ScreenModuleEditorView "PB: KP8 Stop Runtime (Text Label)" 68x66
   Button "Station Select" at 0,0 size 68x66; TextOff 'STOP RUNTIME'
      Appearance <- "Interface.animate"
*)

(* ===== HMI "HMI_RT_1" =====
system functions are stored by id; their names below are inferred from use

ScreenModuleEditorView "PB: Graphic/Text List" 65x45
   Button "Previous Station Group" at 0,0 size 65x45; TextOff 'Text'
      on Press: SetBit("Interface.actuate")
      Visibility <- "Interface.animate"
      ObjectEnable <- "Interface.animate"
      Appearance <- "Interface.animate"
*)

(* ===== HMI "HMI_RT_1" =====
system functions are stored by id; their names below are inferred from use

ScreenModuleEditorView "PB: Static Text Label" 274x45
   Button "Select All Stations" at 0,0 size 274x45; TextOff 'Text'
      on Press: function_b14e0dd5("Interface.actuate", 0)
      Appearance <- "Interface.animate"
*)

(* ===== HMI "HMI_RT_1" =====
system functions are stored by id; their names below are inferred from use

ScreenModuleEditorView "PB: Static Text Label" 274x45
   Button "Select All Stations" at 0,0 size 274x45; TextOff 'Text'
      on Press: function_b14e0dd5("Interface.actuate", 0)
      Appearance <- "Interface.animate"
*)

(* ===== HMI "HMI_RT_1" =====
system functions are stored by id; their names below are inferred from use

ScreenModuleEditorView "PB: Graphic/Text List" 65x45
   Button "Previous Station Group" at 0,0 size 65x45; TextOff 'Text'
      on Press: SetBit("Interface.actuate")
      Visibility <- "Interface.animate"
      ObjectEnable <- "Interface.animate"
      Appearance <- "Interface.animate"
*)

(* ===== HMI "HMI_RT_1" =====
system functions are stored by id; their names below are inferred from use

ScreenModuleEditorView "PB: Station Select (Text Label)" 205x65
   Button "Station Select" at 0,0 size 205x65; TextOff 'Text'
      on Press: function_b14e0dd5("Interface.actuate", 0)
      Appearance <- "Interface.animate"
*)

(* ===== HMI "HMI_RT_1" =====
system functions are stored by id; their names below are inferred from use

ScreenModuleEditorView "PB: Graphic/Text List" 65x45
   Button "Previous Station Group" at 0,0 size 65x45; TextOff 'Text'
      on Press: function_b14e0dd5("Interface.actuate", 0)
      Visibility <- "Interface.animate"
      ObjectEnable <- "Interface.animate"
      Appearance <- "Interface.animate"
*)

(* ===== HMI "HMI_RT_1" =====
system functions are stored by id; their names below are inferred from use

ScreenModuleEditorView "Drop Zone Label" 240x40
   IOField "Drop Zone Entry" at 171,0 size 69x40; FormatPattern ??
      on OnFinishInput: SetBit("Interface.inputFinished")
      Appearance <- "Interface.animate.ioField"
      ObjectEnable <- "Interface.animate.ioField"
      Visibility <- "Interface.animate.ioField"
      ProcessValue <- "Interface.value"
   TextField "Drop Zone Label" at 0,0 size 240x40; Text 'Drop Zone:'
      Visibility <- "Interface.animate.bg"
      Appearance <- "Interface.animate.bg"
*)

(* ===== HMI "HMI_RT_1" =====
system functions are stored by id; their names below are inferred from use

ScreenModuleEditorView "IO Field: Double Width; Stacked" 414x50
   IOField "PN Entry Field" at 0,0 size 414x50; FormatPattern ????????????????????????????????????????
      on OnFinishInput: SetBit("Interface.inputFinished")
      Appearance <- "Interface.animate"
      ObjectEnable <- "Interface.animate"
      ProcessValue <- "Interface.value"
*)

(* ===== HMI "HMI_RT_1" =====
system functions are stored by id; their names below are inferred from use

ScreenModuleEditorView "IO Field: Timer" 137x50
   IOField "Allotted Time Entry Field" at 0,0 size 137x50; FormatPattern ???????
      on OnFinishInput: SetBit("Interface.inputFinished")
      Appearance <- "Interface.animate"
      ObjectEnable <- "Interface.animate"
      ProcessValue <- "Interface.value"
*)

(* ===== HMI "HMI_RT_1" =====

ScreenModuleEditorView "LED Row" 440x28
   TextField "tfLine" at 0,0 size 110x28; Text 'Text'
      Visibility <- "interface.tfLine.visibility"
      Appearance <- "interface.tfLine.animator"
   TextField "tfTime" at 349,0 size 91x28; Text 'Text'
      Visibility <- "interface.tfTime.visibility"
      Appearance <- "interface.tfTime.animator"
   TextField "tfDropZone" at 105,0 size 42x28; Text 'Text'
      Visibility <- "interface.tfDropZone.visibility"
      Appearance <- "interface.tfDropZone.animator"
   TextField "tfSLPartNumber" at 146,0 size 209x28; Text 'Text'
      Visibility <- "interface.tfPartNumber.count"
      Appearance <- "interface.tfPartNumber.animator"
   TextField "tfDLPartNumber" at 146,0 size 209x28; Text 'Text'
      Visibility <- "interface.tfPartNumber.count"
      Appearance <- "interface.tfPartNumber.animator"
*)

(* ===== HMI "HMI_RT_1" =====
system functions are stored by id; their names below are inferred from use

ScreenModuleEditorView "Line Label" 267x40
   IOField "Line" at 86,0 size 181x40; FormatPattern ?????????
      on OnFinishInput: SetBit("interface.inputFinished")
      Appearance <- "interface.animate.ioField"
      ObjectEnable <- "interface.animate.ioField"
      Visibility <- "interface.animate.ioField"
      ProcessValue <- "interface.value"
   TextField "Line Label" at 0,0 size 267x40; Text 'Line:'
      Visibility <- "interface.animate.bg"
      Appearance <- "interface.animate.bg"
*)

(* ===== HMI "HMI_RT_1" =====
system functions are stored by id; their names below are inferred from use

ScreenModuleEditorView "PB: Graphic/Text List" 65x45
   Button "Previous Station Group" at 0,0 size 65x45; TextOff 'Text'
      on Press: function_b14e0dd5("Interface.actuate", 0)
      Visibility <- "Interface.animate"
      ObjectEnable <- "Interface.animate"
      Appearance <- "Interface.animate"
*)

(* ===== HMI "HMI_RT_1" =====
system functions are stored by id; their names below are inferred from use

ScreenModuleEditorView "PB: KP8 Button Select (Text Label)" 68x66
   Button "Station Select" at 0,0 size 68x66; TextOff 'Text'
      on Press: function_b14e0dd5("Interface.actuate", 0)
      Appearance <- "Interface.animate"
*)

(* ===== HMI "HMI_RT_1" =====

ScreenModuleEditorView "PB: KP8 Reset Button (Text Label" 68x66
   Button "Station Select" at 0,0 size 68x66; TextOff 'RESET SELECTED'
      Appearance <- "Interface.animate"
*)

(* ===== HMI "HMI_RT_1" =====

ScreenModuleEditorView "PB: KP8 Stop Runtime (Text Label)" 68x66
   Button "Station Select" at 0,0 size 68x66; TextOff 'STOP RUNTIME'
      Appearance <- "Interface.animate"
*)

(* ===== HMI "HMI_RT_1" =====
system functions are stored by id; their names below are inferred from use

ScreenModuleEditorView "PB: Station Select (Text Label)" 205x65
   Button "Station Select" at 0,0 size 205x65; TextOff 'Text'
      on Press: function_b14e0dd5("Interface.actuate", 0)
      Appearance <- "Interface.animate"
*)

(* ===== HMI "HMI_RT_1" =====
system functions are stored by id; their names below are inferred from use

ScreenModuleEditorView "PB: Static Text Label" 274x45
   Button "Select All Stations" at 0,0 size 274x45; TextOff 'Text'
      on Press: function_b14e0dd5("Interface.actuate", 0)
      Appearance <- "Interface.animate"
*)

(* ===== HMI "HMI_RT_1" =====
system functions are stored by id; their names below are inferred from use

ScreenModuleEditorView "Station Assignment: Button Details" 513x74
   TextField "Button Label" at 0,0 size 75x74; Text 'Text'
      Visibility <- "Interface.label.animate"
      Appearance <- "Interface.label.animate"
   TextField "Critical Time" at 70,37 size 122x37; Text 'Text'
      Visibility <- "Interface.critical.animate"
      Appearance <- "Interface.critical.animate"
   TextField "Alloted Time" at 70,0 size 122x38; Text 'Text'
      Visibility <- "Interface.alloted.animate"
      Appearance <- "Interface.alloted.animate"
   TextField "Part Number" at 185,0 size 328x74; Text 'Text'
      Visibility <- "Interface.partNumber.animate"
      Appearance <- "Interface.partNumber.animate"
   Button "Select PB" at 0,0 size 513x74; TextOff 'Text'
      on Press: function_b14e0dd5("Interface.select.actuate", 0)
      Visibility <- "Interface.select.animate"
      ObjectEnable <- "Interface.select.animate"
*)

(* ===== HMI "HMI_RT_1" =====
system functions are stored by id; their names below are inferred from use

ScreenModuleEditorView "Table Row" 1312x52
   TextField "tfLine" at 5,1 size 216x48; Text 'Text'
      Visibility <- "interface.tfLine.visibility"
      Appearance <- "interface.tfLine.animator"
   TextField "tfTime" at 1085,1 size 222x48; Text 'Text'
      Visibility <- "interface.tfTime.visibility"
      Appearance <- "interface.tfTime.animator"
   TextField "tfDropZone" at 211,1 size 236x48; Text 'Text'
      Visibility <- "interface.tfDropZone.visibility"
      Appearance <- "interface.tfDropZone.animator"
   TextField "tfSLPartNumber" at 445,1 size 650x48; Text 'Text'
      Visibility <- "interface.tfPartNumber.count"
      Appearance <- "interface.tfPartNumber.animator"
   Button "pbSelect" at 0,0 size 1312x52; TextOff 'Text'
      on Release: ResetBit("interface.pbSelection.request")
      on Press: SetBit("interface.pbSelection.request")
      Visibility <- "interface.pbSelection.visibility"
   Rectangle "rtBackground" at 0,0 size 1312x52
      Visibility <- "interface.rtBackground.visibility"
   TextField "tfDLPartNumber" at 445,1 size 650x48; Text 'Text'
      Visibility <- "interface.tfPartNumber.count"
      Appearance <- "interface.tfPartNumber.animator"
*)

(* ===== HMI "HMI_RT_1" =====
system functions are stored by id; their names below are inferred from use

ScreenModuleEditorView "PB: Static Text Label" 274x45
   Button "Select All Stations" at 0,0 size 274x45; TextOff 'Text'
      on Press: function_b14e0dd5("Interface.actuate", 0)
      Appearance <- "Interface.animate"
      ObjectEnable <- "Interface.animate"
*)

(* ===== HMI "HMI_RT_1" =====
system functions are stored by id; their names below are inferred from use

ScreenModuleEditorView "PB: KP8 Button Select (Text Label)" 68x66
   Button "Station Select" at 0,0 size 68x66; TextOff 'Text'
      on Press: function_b14e0dd5("Interface.actuate", 0)
      Appearance <- "Interface.animate"
      ObjectEnable <- "Interface.animate"
*)

(* ===== HMI "HMI_RT_1" =====
system functions are stored by id; their names below are inferred from use

ScreenModuleEditorView "PB: KP8 Reset Button (Text Label" 68x66
   Button "Station Select" at 0,0 size 68x66; TextOff 'RESET SELECTED'
      Appearance <- "Interface.animate"
      on Press: function_b14e0dd5("Interface.actuate", 0)
*)

(* ===== HMI "HMI_RT_1" =====
system functions are stored by id; their names below are inferred from use

ScreenModuleEditorView "Drop Zone Label" 240x40
   IOField "Drop Zone Entry" at 171,0 size 69x40; FormatPattern ??
      on OnFinishInput: SetBit("Interface.inputFinished")
      Appearance <- "Interface.animate.ioField"
      ObjectEnable <- "Interface.animate.ioField"
      ProcessValue <- "Interface.value"
      Visibility <- "Interface.animate.ioField"
   TextField "Drop Zone Label" at 0,0 size 240x40; Text 'Drop Zone:'
      Visibility <- "Interface.animate.bg"
      Appearance <- "Interface.animate.bg"
*)

(* ===== HMI "HMI_RT_1" =====
system functions are stored by id; their names below are inferred from use

ScreenModuleEditorView "Drop Zone Label" 240x40
   IOField "Drop Zone Entry" at 171,0 size 69x40; FormatPattern ??
      on OnFinishInput: SetBit("Interface.inputFinished")
      Appearance <- "Interface.animate.ioField"
      Visibility <- "Interface.animate.ioField"
      ObjectEnable <- "Interface.animate.ioField"
      ProcessValue <- "Interface.value"
   TextField "Drop Zone Label" at 0,0 size 240x40; Text 'Drop Zone:'
      Visibility <- "Interface.animate.bg"
      Appearance <- "Interface.animate.bg"
*)

(* ===== HMI "HMI_RT_1" =====
system functions are stored by id; their names below are inferred from use

ScreenModuleEditorView "IO Field: Double Width; Stacked" 414x50
   IOField "PN Entry Field" at 0,0 size 414x50; FormatPattern ????????????????????????????????????????
      on OnFinishInput: SetBit("Interface.inputFinished")
      Appearance <- "Interface.animate"
      ObjectEnable <- "Interface.animate"
      ProcessValue <- "Interface.value"
      Visibility <- "Interface.animate"
*)

(* ===== HMI "HMI_RT_1" =====
system functions are stored by id; their names below are inferred from use

ScreenModuleEditorView "IO Field: Timer" 137x50
   IOField "Allotted Time Entry Field" at 0,0 size 137x50; FormatPattern ???????
      on OnFinishInput: SetBit("Interface.inputFinished")
      Appearance <- "Interface.animate"
      ObjectEnable <- "Interface.animate"
      ProcessValue <- "Interface.value"
      Visibility <- "Interface.animate"
*)

(* ===== HMI "HMI_RT_1" =====

ScreenModuleEditorView "LED Row" 440x28
   TextField "tfLine" at 0,0 size 110x28; Text 'Text'
      Visibility <- "interface.tfLine.visibility"
      Appearance <- "interface.tfLine.animator"
   TextField "tfTime" at 349,0 size 91x28; Text 'Text'
      Visibility <- "interface.tfTime.visibility"
      Appearance <- "interface.tfTime.animator"
   TextField "tfDropZone" at 105,0 size 42x28; Text 'Text'
      Visibility <- "interface.tfDropZone.visibility"
      Appearance <- "interface.tfDropZone.animator"
   TextField "tfSLPartNumber" at 146,0 size 209x28; Text 'Text'
      Visibility <- "interface.tfPartNumber.count"
      Appearance <- "interface.tfPartNumber.animator"
   TextField "tfDLPartNumber" at 146,0 size 209x28; Text 'Text'
      Visibility <- "interface.tfPartNumber.count"
      Appearance <- "interface.tfPartNumber.animator"
*)

(* ===== HMI "HMI_RT_1" =====
system functions are stored by id; their names below are inferred from use

ScreenModuleEditorView "Line Label" 267x40
   IOField "Line" at 86,0 size 181x40; FormatPattern ?????????
      on OnFinishInput: SetBit("interface.inputFinished")
      Appearance <- "interface.animate.ioField"
      ObjectEnable <- "interface.animate.ioField"
      ProcessValue <- "interface.value"
      Visibility <- "interface.animate.ioField"
   TextField "Line Label" at 0,0 size 267x40; Text 'Line:'
      Visibility <- "interface.animate.bg"
      Appearance <- "interface.animate.bg"
*)

(* ===== HMI "HMI_RT_1" =====
system functions are stored by id; their names below are inferred from use

ScreenModuleEditorView "PB: Graphic/Text List" 65x45
   Button "Previous Station Group" at 0,0 size 65x45; TextOff 'Text'
      on Press: function_b14e0dd5("Interface.actuate", 0)
      Visibility <- "Interface.animate"
      ObjectEnable <- "Interface.animate"
      Appearance <- "Interface.animate"
*)

(* ===== HMI "HMI_RT_1" =====
system functions are stored by id; their names below are inferred from use

ScreenModuleEditorView "PB: KP8 Button Select (Text Label)" 68x66
   Button "Station Select" at 0,0 size 68x66; TextOff 'Text'
      on Press: function_b14e0dd5("Interface.actuate", 0)
      Appearance <- "Interface.animate"
      ObjectEnable <- "Interface.animate"
      Visibility <- "Interface.animate"
*)

(* ===== HMI "HMI_RT_1" =====
system functions are stored by id; their names below are inferred from use

ScreenModuleEditorView "PB: KP8 Reset Button (Text Label" 68x66
   Button "Station Select" at 0,0 size 68x66; TextOff 'RESET SELECTED'
      on Press: function_b14e0dd5("Interface.actuate", 0)
      Appearance <- "Interface.animate"
      ObjectEnable <- "Interface.animate"
      Visibility <- "Interface.animate"
*)

(* ===== HMI "HMI_RT_1" =====

ScreenModuleEditorView "PB: KP8 Stop Runtime (Text Label)" 68x66
   Button "Station Select" at 0,0 size 68x66; TextOff 'STOP RUNTIME'
      Appearance <- "Interface.animate"
      ObjectEnable <- "Interface.animate"
      Visibility <- "Interface.animate"
*)

(* ===== HMI "HMI_RT_1" =====
system functions are stored by id; their names below are inferred from use

ScreenModuleEditorView "PB: Station Select (Text Label)" 205x65
   Button "Station Select" at 0,0 size 205x65; TextOff 'Text'
      on Press: function_b14e0dd5("Interface.actuate", 0)
      Appearance <- "Interface.animate"
      ObjectEnable <- "Interface.animate"
      Visibility <- "Interface.animate"
*)

(* ===== HMI "HMI_RT_1" =====
system functions are stored by id; their names below are inferred from use

ScreenModuleEditorView "PB: Static Text Label" 274x45
   Button "Select All Stations" at 0,0 size 274x45; TextOff 'Text'
      on Press: function_b14e0dd5("Interface.actuate", 0)
      Appearance <- "Interface.animate"
      ObjectEnable <- "Interface.animate"
      Visibility <- "Interface.animate"
*)

(* ===== HMI "HMI_RT_1" =====
system functions are stored by id; their names below are inferred from use

ScreenModuleEditorView "Station Assignment: Button Details" 513x74
   TextField "Button Label" at 0,0 size 75x74; Text 'Text'
      Visibility <- "Interface.label.animate"
      Appearance <- "Interface.label.animate"
   TextField "Critical Time" at 70,37 size 122x37; Text 'Text'
      Visibility <- "Interface.critical.animate"
      Appearance <- "Interface.critical.animate"
   TextField "Alloted Time" at 70,0 size 122x38; Text 'Text'
      Visibility <- "Interface.alloted.animate"
      Appearance <- "Interface.alloted.animate"
   TextField "Part Number" at 185,0 size 328x74; Text 'Text'
      Visibility <- "Interface.partNumber.animate"
      Appearance <- "Interface.partNumber.animate"
   Button "Select PB" at 0,0 size 513x74; TextOff 'Text'
      on Press: function_b14e0dd5("Interface.select.actuate", 0)
      Visibility <- "Interface.select.animate"
      ObjectEnable <- "Interface.select.animate"
*)

(* ===== HMI "HMI_RT_1" =====
system functions are stored by id; their names below are inferred from use

ScreenModuleEditorView "Table Row" 1312x52
   TextField "tfLine" at 5,1 size 216x48; Text 'Text'
      Visibility <- "interface.tfLine.animate"
      Appearance <- "interface.tfLine.animate"
   TextField "tfTime" at 1085,1 size 222x48; Text 'Text'
      Appearance <- "interface.tfTime.animate"
      Visibility <- "interface.tfTime.animate"
   TextField "tfDropZone" at 211,1 size 236x48; Text 'Text'
      Visibility <- "interface.tfDropZone.animate"
      Appearance <- "interface.tfDropZone.animate"
   TextField "tfSLPartNumber" at 445,1 size 650x48; Text 'Text'
      Appearance <- "interface.tfPartNumber.animate"
      Visibility <- "interface.tfPartNumber.animate"
   Button "pbSelect" at 0,0 size 1312x52; TextOff 'Text'
      on Press: function_b14e0dd5("interface.pbSelection.actuate", 0)
      Appearance <- "interface.pbSelection.animate"
      ObjectEnable <- "interface.pbSelection.animate"
      Visibility <- "interface.pbSelection.animate"
   Rectangle "rtBackground" at 0,0 size 1312x52
      Appearance <- "interface.rtBackground.animate"
      Visibility <- "interface.rtBackground.animate"
   TextField "tfDLPartNumber" at 445,1 size 650x48; Text 'Text'
      Visibility <- "interface.tfPartNumber.animate"
      Appearance <- "interface.tfPartNumber.animate"
*)

(* ===== HMI "HMI_RT_1" =====
system functions are stored by id; their names below are inferred from use

ScreenModuleEditorView "Table Row" 1312x52
   TextField "tfLine" at 5,1 size 216x48; Text 'Text'
      Visibility <- "interface.tfLine.animate"
      Appearance <- "interface.tfLine.animate"
   TextField "tfTime" at 1085,1 size 222x48; Text 'Text'
      Visibility <- "interface.tfTime.animate"
      Appearance <- "interface.tfTime.animate"
   TextField "tfDropZone" at 211,1 size 236x48; Text 'Text'
      Visibility <- "interface.tfDropZone.animate"
      Appearance <- "interface.tfDropZone.animate"
   TextField "tfSLPartNumber" at 445,1 size 650x48; Text 'Text'
      Visibility <- "interface.tfPartNumber.animate"
      Appearance <- "interface.tfPartNumber.animate"
   Button "pbSelect" at 0,0 size 1312x52; TextOff 'Text'
      on Press: function_b14e0dd5("interface.pbSelection.actuate", 0)
      Appearance <- "interface.pbSelection.animate"
      ObjectEnable <- "interface.pbSelection.animate"
      Visibility <- "interface.pbSelection.animate"
   Rectangle "rtBackground" at 0,0 size 1312x52
      Visibility <- "interface.rtBackground.animate"
      Appearance <- "interface.rtBackground.animate"
   TextField "tfDLPartNumber" at 445,1 size 650x48; Text 'Text'
      Visibility <- "interface.tfPartNumber.animate"
      Appearance <- "interface.tfPartNumber.animate"
*)

(* ===== HMI "HMI_RT_1" =====
system functions are stored by id; their names below are inferred from use

ScreenModuleEditorView "Table Row" 1312x52
   TextField "tfLine" at 5,1 size 216x48; Text 'Text'
      Visibility <- "interface.tfLine.animate"
      Appearance <- "interface.tfLine.animate"
   TextField "tfTime" at 1085,1 size 222x48; Text 'Text'
      Visibility <- "interface.tfTime.animate"
      Appearance <- "interface.tfTime.animate"
   TextField "tfDropZone" at 211,1 size 236x48; Text 'Text'
      Visibility <- "interface.tfDropZone.animate"
      Appearance <- "interface.tfDropZone.animate"
   TextField "tfSLPartNumber" at 445,1 size 650x48; Text 'Text'
      Appearance <- "interface.tfPartNumber.animateSL"
      Visibility <- "interface.tfPartNumber.animateDL"
   Button "pbSelect" at 0,0 size 1312x52; TextOff 'Text'
      on Press: function_b14e0dd5("interface.pbSelection.actuate", 0)
      Appearance <- "interface.pbSelection.animate"
      ObjectEnable <- "interface.pbSelection.animate"
      Visibility <- "interface.pbSelection.animate"
   Rectangle "rtBackground" at 0,0 size 1312x52
      Visibility <- "interface.rtBackground.animate"
      Appearance <- "interface.rtBackground.animate"
   TextField "tfDLPartNumber" at 445,1 size 650x48; Text 'Text'
      Appearance <- "interface.tfPartNumber.animateDL"
      Visibility <- "interface.tfPartNumber.animateDL"
*)

(* ===== HMI "HMI_RT_1" =====
system functions are stored by id; their names below are inferred from use

ScreenModuleEditorView "Table Row" 1312x52
   TextField "tfLine" at 5,1 size 216x48; Text 'Text'
      Visibility <- "interface.tfLine.animate"
      Appearance <- "interface.tfLine.animate"
   TextField "tfTime" at 1085,1 size 222x48; Text 'Text'
      Visibility <- "interface.tfTime.animate"
      Appearance <- "interface.tfTime.animate"
   TextField "tfDropZone" at 211,1 size 236x48; Text 'Text'
      Visibility <- "interface.tfDropZone.animate"
      Appearance <- "interface.tfDropZone.animate"
   TextField "tfSLPartNumber" at 445,1 size 650x48; Text 'Text'
      Visibility <- "interface.tfPartNumber.animateDL"
      Appearance <- "interface.tfPartNumber.animateSL"
   Button "pbSelect" at 0,0 size 1312x52; TextOff 'Text'
      on Press: function_b14e0dd5("interface.pbSelection.actuate", 0)
      Appearance <- "interface.pbSelection.animate"
      ObjectEnable <- "interface.pbSelection.animate"
      Visibility <- "interface.pbSelection.animate"
   Rectangle "rtBackground" at 0,0 size 1312x52
      Visibility <- "interface.rtBackground.animate"
      Appearance <- "interface.rtBackground.animate"
   TextField "tfDLPartNumber" at 445,1 size 650x48; Text 'Text'
      Visibility <- "interface.tfPartNumber.animateDL"
      Appearance <- "interface.tfPartNumber.animateDL"
*)

(* ===== HMI "HMI_RT_1" =====
system functions are stored by id; their names below are inferred from use

ScreenModuleEditorView "Table Row" 1312x52
   TextField "tfLine" at 5,1 size 216x48; Text 'Text'
      Visibility <- "interface.tfLine.animate"
      Appearance <- "interface.tfLine.animate"
   TextField "tfTime" at 1085,1 size 222x48; Text 'Text'
      Visibility <- "interface.tfTime.animate"
      Appearance <- "interface.tfTime.animate"
   TextField "tfDropZone" at 211,1 size 236x48; Text 'Text'
      Visibility <- "interface.tfDropZone.animate"
      Appearance <- "interface.tfDropZone.animate"
   TextField "tfSLPartNumber" at 445,1 size 650x48; Text 'Text'
      Appearance <- "interface.tfPartNumber.animateSL"
      Visibility <- "interface.tfPartNumber.animateSL"
   Button "pbSelect" at 0,0 size 1312x52; TextOff 'Text'
      on Press: function_b14e0dd5("interface.pbSelection.actuate", 0)
      Appearance <- "interface.pbSelection.animate"
      ObjectEnable <- "interface.pbSelection.animate"
      Visibility <- "interface.pbSelection.animate"
   Rectangle "rtBackground" at 0,0 size 1312x52
      Visibility <- "interface.rtBackground.animate"
      Appearance <- "interface.rtBackground.animate"
   TextField "tfDLPartNumber" at 445,1 size 650x48; Text 'Text'
      Visibility <- "interface.tfPartNumber.animateDL"
      Appearance <- "interface.tfPartNumber.animateDL"
*)

(* ===== HMI "HMI_RT_1" =====

ScreenModuleEditorView "LED Row" 440x28
   TextField "tfLine" at 0,0 size 110x28; Text 'Text'
      Appearance <- "interface.tfLine.animate"
      Visibility <- "interface.tfLine.animate"
   TextField "tfTime" at 349,0 size 91x28; Text 'Text'
      Visibility <- "interface.tfTime.animate"
      Appearance <- "interface.tfTime.animate"
   TextField "tfDropZone" at 105,0 size 42x28; Text 'Text'
      Appearance <- "interface.tfDropZone.animate"
      Visibility <- "interface.tfDropZone.animate"
   TextField "tfSLPartNumber" at 146,0 size 209x28; Text 'Text'
      Visibility <- "interface.tfPartNumber.animateSL"
      Appearance <- "interface.tfPartNumber.animateSL"
   TextField "tfDLPartNumber" at 146,0 size 209x28; Text 'Text'
      Appearance <- "interface.tfPartNumber.animateDL"
      Visibility <- "interface.tfPartNumber.animateDL"
*)

(* ===== HMI "HMI_RT_1" =====
system functions are stored by id; their names below are inferred from use

ScreenModuleEditorView "Table Row" 1312x52
   TextField "tfLine" at 5,1 size 216x48; Text 'Text'
      Visibility <- "interface.tfLine.animate"
      Appearance <- "interface.tfLine.animate"
   TextField "tfTime" at 1085,1 size 222x48; Text 'Text'
      Visibility <- "interface.tfTime.animate"
      Appearance <- "interface.tfTime.animate"
   TextField "tfDropZone" at 211,1 size 236x48; Text 'Text'
      Visibility <- "interface.tfDropZone.animate"
      Appearance <- "interface.tfDropZone.animate"
   TextField "tfSLPartNumber" at 445,1 size 650x48; Text 'Text'
      Visibility <- "interface.tfPartNumber.animateSL"
      Appearance <- "interface.tfPartNumber.animateSL"
   Button "pbSelect" at 0,0 size 1312x52; TextOff 'Text'
      on Press: function_b14e0dd5("interface.pbSelection.actuate", 0)
      Appearance <- "interface.pbSelection.animate"
      ObjectEnable <- "interface.pbSelection.animate"
      Visibility <- "interface.pbSelection.animate"
   Rectangle "rtBackground" at 0,0 size 1312x52
      Visibility <- "interface.rtBackground.animate"
      Appearance <- "interface.rtBackground.animate"
   TextField "tfDLPartNumber" at 445,1 size 650x48; Text 'Text'
      Visibility <- "interface.tfPartNumber.animateDL"
      Appearance <- "interface.tfPartNumber.animateDL"
*)

(* ===== HMI "HMI_RT_1" =====

ScreenModuleEditorView "LED Row" 440x28
   TextField "tfLine" at 0,0 size 110x28; Text 'Text'
      Visibility <- "interface.tfLine.animate"
      Appearance <- "interface.tfLine.animate"
   TextField "tfTime" at 349,0 size 91x28; Text 'Text'
      Visibility <- "interface.tfTime.animate"
      Appearance <- "interface.tfTime.animate"
   TextField "tfDropZone" at 105,0 size 42x28; Text 'Text'
      Visibility <- "interface.tfDropZone.animate"
      Appearance <- "interface.tfDropZone.animate"
   TextField "tfSLPartNumber" at 146,0 size 209x28; Text 'Text'
      Visibility <- "interface.tfPartNumber.animateSL"
      Appearance <- "interface.tfPartNumber.animateSL"
   TextField "tfDLPartNumber" at 146,0 size 209x28; Text 'Text'
      Visibility <- "interface.tfPartNumber.animateDL"
      Appearance <- "interface.tfPartNumber.animateDL"
*)

(* ===== HMI "HMI_RT_1" =====
system functions are stored by id; their names below are inferred from use

ScreenModuleEditorView "Table Row" 1312x52
   TextField "tfLine" at 5,1 size 216x48; Text 'Text'
      Visibility <- "interface.tfLine.animate"
      Appearance <- "interface.tfLine.animate"
   TextField "tfTime" at 1085,1 size 222x48; Text 'Text'
      Visibility <- "interface.tfTime.animate"
      Appearance <- "interface.tfTime.animate"
   TextField "tfDropZone" at 211,1 size 236x48; Text 'Text'
      Visibility <- "interface.tfDropZone.animate"
      Appearance <- "interface.tfDropZone.animate"
   TextField "tfSLPartNumber" at 445,1 size 650x48; Text 'Text'
      Visibility <- "interface.tfPartNumber.animateSL"
      Appearance <- "interface.tfPartNumber.animateSL"
   Button "pbSelect" at 0,0 size 1312x52; TextOff 'Text'
      on Press: SetBit("interface.pbSelection.actuate")
      Appearance <- "interface.pbSelection.animate"
      ObjectEnable <- "interface.pbSelection.animate"
      Visibility <- "interface.pbSelection.animate"
      on Release: ResetBit("interface.pbSelection.actuate")
   Rectangle "rtBackground" at 0,0 size 1312x52
      Visibility <- "interface.rtBackground.animate"
      Appearance <- "interface.rtBackground.animate"
   TextField "tfDLPartNumber" at 445,1 size 650x48; Text 'Text'
      Visibility <- "interface.tfPartNumber.animateDL"
      Appearance <- "interface.tfPartNumber.animateDL"
*)

(* ===== HMI "HMI_RT_1" =====
system functions are stored by id; their names below are inferred from use

ScreenModuleEditorView "Table Row" 1312x52
   TextField "tfLine" at 5,1 size 216x48; Text 'Text'
      Visibility <- "interface.tfLine.animate"
      Appearance <- "interface.tfLine.animate"
   TextField "tfTime" at 1085,1 size 222x48; Text 'Text'
      Visibility <- "interface.tfTime.animate"
      Appearance <- "interface.tfTime.animate"
   TextField "tfDropZone" at 211,1 size 236x48; Text 'Text'
      Visibility <- "interface.tfDropZone.animate"
      Appearance <- "interface.tfDropZone.animate"
   TextField "tfSLPartNumber" at 445,1 size 650x48; Text 'Text'
      Visibility <- "interface.tfPartNumber.animateSL"
      Appearance <- "interface.tfPartNumber.animateSL"
   Button "pbSelect" at 0,0 size 1312x52; TextOff 'Text'
      on Press: function_b14e0dd5("interface.pbSelection.actuate", 0)
      Appearance <- "interface.pbSelection.animate"
      ObjectEnable <- "interface.pbSelection.animate"
      Visibility <- "interface.pbSelection.animate"
   Rectangle "rtBackground" at 0,0 size 1312x52
      Visibility <- "interface.rtBackground.animate"
      Appearance <- "interface.rtBackground.animate"
   TextField "tfDLPartNumber" at 445,1 size 650x48; Text 'Text'
      Visibility <- "interface.tfPartNumber.animateDL"
      Appearance <- "interface.tfPartNumber.animateDL"
*)

(* ===== HMI "HMI_RT_1" =====
system functions are stored by id; their names below are inferred from use

ScreenModuleEditorView "PB: Graphic/Text List" 65x45
   Button "Previous Station Group" at 0,0 size 65x45; TextOff 'Text'
      on Press: function_b14e0dd5("Interface.actuate", 0)
      Visibility <- "Interface.animate"
      ObjectEnable <- "Interface.animate"
      Appearance <- "Interface.animate"
*)

(* ===== HMI "HMI_RT_1" =====
system functions are stored by id; their names below are inferred from use

ScreenModuleEditorView "PB: Graphic/Text List" 65x45
   Button "Previous Station Group" at 0,0 size 65x45; TextOff 'Text'
      on Press: function_b14e0dd5("Interface.actuate", 0)
      Visibility <- "Interface.animate"
      ObjectEnable <- "Interface.animate"
      Appearance <- "Interface.animate"
*)

(* ===== HMI "HMI_RT_1" =====
system functions are stored by id; their names below are inferred from use

ScreenModuleEditorView "Table Row" 1312x52
   TextField "tfLine" at 5,1 size 216x48; Text 'Text'
      Visibility <- "interface.tfLine.animate"
      Appearance <- "interface.tfLine.animate"
   TextField "tfTime" at 1085,1 size 222x48; Text 'Text'
      Visibility <- "interface.tfTime.animate"
      Appearance <- "interface.tfTime.animate"
   TextField "tfDropZone" at 211,1 size 236x48; Text 'Text'
      Visibility <- "interface.tfDropZone.animate"
      Appearance <- "interface.tfDropZone.animate"
   TextField "tfSLPartNumber" at 445,1 size 650x48; Text 'Text'
      Visibility <- "interface.tfPartNumber.animateSL"
      Appearance <- "interface.tfPartNumber.animateSL"
   Button "pbSelect" at 0,0 size 1312x52; TextOff 'Text'
      on Press: SetBit("interface.pbSelection.actuate")
      Appearance <- "interface.pbSelection.animate"
      ObjectEnable <- "interface.pbSelection.animate"
      Visibility <- "interface.pbSelection.animate"
      on Release: ResetBit("interface.pbSelection.actuate")
   Rectangle "rtBackground" at 0,0 size 1312x52
      Visibility <- "interface.rtBackground.animate"
      Appearance <- "interface.rtBackground.animate"
   TextField "tfDLPartNumber" at 445,1 size 650x48; Text 'Text'
      Visibility <- "interface.tfPartNumber.animateDL"
      Appearance <- "interface.tfPartNumber.animateDL"
*)

(* ===== HMI "HMI_RT_1" =====
system functions are stored by id; their names below are inferred from use

ScreenModuleEditorView "Station Sim" 102x228
   TextField "Station Label" at 0,0 size 102x20; Text 'Text'
      Appearance <- "Interface.stn.animate"
   Button "B7" at 0,22 size 50x50; TextOff 'Text'
      Appearance <- "Interface.btn.animate[7]"
      on Press: function_b14e0dd5("Interface.btn.actuate", 7)
   Button "B6" at 0,74 size 50x50; TextOff 'Text'
      Appearance <- "Interface.btn.animate[6]"
      on Press: function_b14e0dd5("Interface.btn.actuate", 6)
   Button "B5" at 0,126 size 50x50; TextOff 'Text'
      Appearance <- "Interface.btn.animate[5]"
      on Press: function_b14e0dd5("Interface.btn.actuate", 5)
   Button "B4" at 0,178 size 50x50; TextOff 'Text'
      Appearance <- "Interface.btn.animate[4]"
      on Press: function_b14e0dd5("Interface.btn.actuate", 4)
   Button "B3" at 52,22 size 50x50; TextOff 'Text'
      Appearance <- "Interface.btn.animate[3]"
      on Press: function_b14e0dd5("Interface.btn.actuate", 3)
   Button "B2" at 52,74 size 50x50; TextOff 'Text'
      Appearance <- "Interface.btn.animate[2]"
      on Press: function_b14e0dd5("Interface.btn.actuate", 2)
   Button "B1" at 52,126 size 50x50; TextOff 'Text'
      Appearance <- "Interface.btn.animate[1]"
      on Press: function_b14e0dd5("Interface.btn.actuate", 1)
   Button "B0" at 52,178 size 50x50; TextOff 'Text'
      Appearance <- "Interface.btn.animate[0]"
      on Press: function_b14e0dd5("Interface.btn.actuate", 0)
*)

(* ===== HMI "HMI_RT_1" =====
system functions are stored by id; their names below are inferred from use

ScreenModuleEditorView "Station Sim" 102x228
   TextField "Station Label" at 0,0 size 102x20; Text 'Text'
      Appearance <- "Interface.stn.animate"
   Button "B7" at 0,22 size 50x50; TextOff 'Text'
      on Press: function_b14e0dd5("Interface.btn.actuate", 7)
      Appearance <- "Interface.btn.animate[7]"
   Button "B6" at 0,74 size 50x50; TextOff 'Text'
      on Press: function_b14e0dd5("Interface.btn.actuate", 6)
      Appearance <- "Interface.btn.animate[6]"
   Button "B5" at 0,126 size 50x50; TextOff 'Text'
      on Press: function_b14e0dd5("Interface.btn.actuate", 5)
      Appearance <- "Interface.btn.animate[5]"
   Button "B4" at 0,178 size 50x50; TextOff 'Text'
      on Press: function_b14e0dd5("Interface.btn.actuate", 4)
      Appearance <- "Interface.btn.animate[4]"
   Button "B3" at 52,22 size 50x50; TextOff 'Text'
      on Press: function_b14e0dd5("Interface.btn.actuate", 3)
      Appearance <- "Interface.btn.animate[3]"
   Button "B2" at 52,74 size 50x50; TextOff 'Text'
      on Press: function_b14e0dd5("Interface.btn.actuate", 2)
      Appearance <- "Interface.btn.animate[2]"
   Button "B1" at 52,126 size 50x50; TextOff 'Text'
      on Press: function_b14e0dd5("Interface.btn.actuate", 1)
      Appearance <- "Interface.btn.animate[1]"
   Button "B0" at 52,178 size 50x50; TextOff 'Text'
      on Press: function_b14e0dd5("Interface.btn.actuate", 0)
      Appearance <- "Interface.btn.animate[0]"
*)

(* ===== HMI "HMI_RT_1" =====
system functions are stored by id; their names below are inferred from use

ScreenModuleEditorView "Station Sim" 106x232
   TextField "Station Label" at 2,2 size 102x20; Text 'Text'
      Appearance <- "Interface.stn.animate"
   Button "B7" at 2,24 size 50x50; TextOff 'Text'
      on Press: function_b14e0dd5("Interface.btn.actuate", 7)
      Appearance <- "Interface.btn.animate[7]"
   Button "B6" at 2,76 size 50x50; TextOff 'Text'
      on Press: function_b14e0dd5("Interface.btn.actuate", 6)
      Appearance <- "Interface.btn.animate[6]"
   Button "B5" at 2,128 size 50x50; TextOff 'Text'
      on Press: function_b14e0dd5("Interface.btn.actuate", 5)
      Appearance <- "Interface.btn.animate[5]"
   Button "B4" at 2,180 size 50x50; TextOff 'Text'
      on Press: function_b14e0dd5("Interface.btn.actuate", 4)
      Appearance <- "Interface.btn.animate[4]"
   Button "B3" at 54,24 size 50x50; TextOff 'Text'
      on Press: function_b14e0dd5("Interface.btn.actuate", 3)
      Appearance <- "Interface.btn.animate[3]"
   Button "B2" at 54,76 size 50x50; TextOff 'Text'
      on Press: function_b14e0dd5("Interface.btn.actuate", 2)
      Appearance <- "Interface.btn.animate[2]"
   Button "B1" at 54,128 size 50x50; TextOff 'Text'
      on Press: function_b14e0dd5("Interface.btn.actuate", 1)
      Appearance <- "Interface.btn.animate[1]"
   Button "B0" at 54,180 size 50x50; TextOff 'Text'
      on Press: function_b14e0dd5("Interface.btn.actuate", 0)
      Appearance <- "Interface.btn.animate[0]"
*)

(* ===== HMI "HMI_RT_1" =====
system functions are stored by id; their names below are inferred from use

ScreenModuleEditorView "Station Sim" 106x232
   Button "B7" at 3,26 size 48x48; TextOff 'Text'
      on Press: function_b14e0dd5("Interface.btn.actuate", 7)
      Appearance <- "Interface.btn.animate[7]"
   Button "B3" at 54,26 size 48x48; TextOff 'Text'
      on Press: function_b14e0dd5("Interface.btn.actuate", 3)
      Appearance <- "Interface.btn.animate[3]"
   Button "B6" at 3,77 size 48x48; TextOff 'Text'
      on Press: function_b14e0dd5("Interface.btn.actuate", 6)
      Appearance <- "Interface.btn.animate[6]"
   Button "B2" at 54,77 size 48x48; TextOff 'Text'
      on Press: function_b14e0dd5("Interface.btn.actuate", 2)
      Appearance <- "Interface.btn.animate[2]"
   Button "B5" at 3,128 size 48x48; TextOff 'Text'
      on Press: function_b14e0dd5("Interface.btn.actuate", 5)
      Appearance <- "Interface.btn.animate[5]"
   Button "B1" at 54,128 size 48x48; TextOff 'Text'
      on Press: function_b14e0dd5("Interface.btn.actuate", 1)
      Appearance <- "Interface.btn.animate[1]"
   Button "B4" at 3,179 size 48x48; TextOff 'Text'
      on Press: function_b14e0dd5("Interface.btn.actuate", 4)
      Appearance <- "Interface.btn.animate[4]"
   Button "B0" at 54,179 size 48x48; TextOff 'Text'
      on Press: function_b14e0dd5("Interface.btn.actuate", 0)
      Appearance <- "Interface.btn.animate[0]"
   TextField "Station Label" at 1,1 size 104x21; Text 'Text'
      Appearance <- "Interface.stn.animate"
*)

(* ===== HMI "HMI_RT_1" =====
system functions are stored by id; their names below are inferred from use

ScreenModuleEditorView "Station Sim" 106x232
   Button "B7" at 3,26 size 48x48; TextOff 'Text'
      on Press: function_b14e0dd5("Interface.btn.actuate", 7)
      Appearance <- "Interface.btn.animate[7]"
   Button "B3" at 54,26 size 48x48; TextOff 'Text'
      on Press: function_b14e0dd5("Interface.btn.actuate", 3)
      Appearance <- "Interface.btn.animate[3]"
   Button "B6" at 3,77 size 48x48; TextOff 'Text'
      on Press: function_b14e0dd5("Interface.btn.actuate", 6)
      Appearance <- "Interface.btn.animate[6]"
   Button "B2" at 54,77 size 48x48; TextOff 'Text'
      on Press: function_b14e0dd5("Interface.btn.actuate", 2)
      Appearance <- "Interface.btn.animate[2]"
   Button "B5" at 3,128 size 48x48; TextOff 'Text'
      on Press: function_b14e0dd5("Interface.btn.actuate", 5)
      Appearance <- "Interface.btn.animate[5]"
   Button "B1" at 54,128 size 48x48; TextOff 'Text'
      on Press: function_b14e0dd5("Interface.btn.actuate", 1)
      Appearance <- "Interface.btn.animate[1]"
   Button "B4" at 3,179 size 48x48; TextOff 'Text'
      on Press: function_b14e0dd5("Interface.btn.actuate", 4)
      Appearance <- "Interface.btn.animate[4]"
   Button "B0" at 54,179 size 48x48; TextOff 'Text'
      on Press: function_b14e0dd5("Interface.btn.actuate", 0)
      Appearance <- "Interface.btn.animate[0]"
   TextField "Station Label" at 1,1 size 104x21; Text 'Text'
      Appearance <- "Interface.stn.animate"
*)

(* ===== HMI "HMI_RT_1" =====
system functions are stored by id; their names below are inferred from use

ScreenModuleEditorView "Table Row" 1312x52
   TextField "tfLine" at 5,1 size 216x48; Text 'Text'
      Visibility <- "interface.tfLine.animate"
      Appearance <- "interface.tfLine.animate"
   TextField "tfTime" at 1085,1 size 222x48; Text 'Text'
      Visibility <- "interface.tfTime.animate"
      Appearance <- "interface.tfTime.animate"
   TextField "tfDropZone" at 211,1 size 236x48; Text 'Text'
      Visibility <- "interface.tfDropZone.animate"
      Appearance <- "interface.tfDropZone.animate"
   TextField "tfSLPartNumber" at 445,1 size 650x48; Text 'Text'
      Visibility <- "interface.tfPartNumber.animateSL"
      Appearance <- "interface.tfPartNumber.animateSL"
   Button "pbSelect" at 0,0 size 1312x52; TextOff 'Text'
      on Release: ResetBit("interface.pbSelection.actuate")
      on Press: SetBit("interface.pbSelection.actuate")
      Appearance <- "interface.pbSelection.animate"
      ObjectEnable <- "interface.pbSelection.animate"
      Visibility <- "interface.pbSelection.animate"
   Rectangle "rtBackground" at 0,0 size 1312x52
      Visibility <- "interface.rtBackground.animate"
      Appearance <- "interface.rtBackground.animate"
   TextField "tfDLPartNumber" at 445,1 size 650x48; Text 'Text'
      Visibility <- "interface.tfPartNumber.animateDL"
      Appearance <- "interface.tfPartNumber.animateDL"
*)

(* ===== HMI "HMI_RT_1" =====
system functions are stored by id; their names below are inferred from use

ScreenModuleEditorView "Station Assignment: Button Details" 513x74
   TextField "Button Label" at 0,0 size 75x74; Text 'Text'
      Visibility <- "Interface.label.animate"
      Appearance <- "Interface.label.animate"
   TextField "Critical Time" at 70,37 size 122x37; Text 'Text'
      Visibility <- "Interface.critical.animate"
      Appearance <- "Interface.critical.animate"
   TextField "Alloted Time" at 70,0 size 122x38; Text 'Text'
      Visibility <- "Interface.alloted.animate"
      Appearance <- "Interface.alloted.animate"
   TextField "Part Number" at 185,0 size 328x74; Text 'Text'
      Visibility <- "Interface.partNumber.animate"
      Appearance <- "Interface.partNumber.animate"
   Button "Select PB" at 0,0 size 513x74; TextOff 'Text'
      on Press: function_b14e0dd5("Interface.select.actuate", 0)
      Visibility <- "Interface.select.animate"
      ObjectEnable <- "Interface.select.animate"
*)

(* ===== HMI "HMI_RT_1" =====
system functions are stored by id; their names below are inferred from use

ScreenModuleEditorView "PB: Static Text Label" 274x45
   Button "Select All Stations" at 0,0 size 274x45; TextOff 'Text'
      on Press: function_b14e0dd5("Interface.actuate", 0)
      Appearance <- "Interface.animate"
      ObjectEnable <- "Interface.animate"
      Visibility <- "Interface.animate"
*)

(* ===== HMI "HMI_RT_1" =====
system functions are stored by id; their names below are inferred from use

ScreenModuleEditorView "PB: Station Select (Text Label)" 205x65
   Button "Station Select" at 0,0 size 205x65; TextOff 'Text'
      on Press: function_b14e0dd5("Interface.actuate", 0)
      Appearance <- "Interface.animate"
      ObjectEnable <- "Interface.animate"
      Visibility <- "Interface.animate"
*)

(* ===== HMI "HMI_RT_1" =====

ScreenModuleEditorView "PB: KP8 Stop Runtime (Text Label)" 68x66
   Button "Station Select" at 0,0 size 68x66; TextOff 'STOP RUNTIME'
      Appearance <- "Interface.animate"
      ObjectEnable <- "Interface.animate"
      Visibility <- "Interface.animate"
*)

(* ===== HMI "HMI_RT_1" =====
system functions are stored by id; their names below are inferred from use

ScreenModuleEditorView "PB: KP8 Reset Button (Text Label" 68x66
   Button "Station Select" at 0,0 size 68x66; TextOff 'RESET SELECTED'
      on Press: function_b14e0dd5("Interface.actuate", 0)
      Appearance <- "Interface.animate"
      ObjectEnable <- "Interface.animate"
      Visibility <- "Interface.animate"
*)

(* ===== HMI "HMI_RT_1" =====
system functions are stored by id; their names below are inferred from use

ScreenModuleEditorView "PB: KP8 Button Select (Text Label)" 68x66
   Button "Station Select" at 0,0 size 68x66; TextOff 'Text'
      on Press: function_b14e0dd5("Interface.actuate", 0)
      Appearance <- "Interface.animate"
      ObjectEnable <- "Interface.animate"
      Visibility <- "Interface.animate"
*)

(* ===== HMI "HMI_RT_1" =====
system functions are stored by id; their names below are inferred from use

ScreenModuleEditorView "PB: Graphic/Text List" 65x45
   Button "Previous Station Group" at 0,0 size 65x45; TextOff 'Text'
      on Press: function_b14e0dd5("Interface.actuate", 0)
      Visibility <- "Interface.animate"
      ObjectEnable <- "Interface.animate"
      Appearance <- "Interface.animate"
*)

(* ===== HMI "HMI_RT_1" =====
system functions are stored by id; their names below are inferred from use

ScreenModuleEditorView "Line Label" 267x40
   IOField "Line" at 86,0 size 181x40; FormatPattern ?????????
      on OnFinishInput: SetBit("interface.inputFinished")
      Appearance <- "interface.animate.ioField"
      Visibility <- "interface.animate.ioField"
      ObjectEnable <- "interface.animate.ioField"
      ProcessValue <- "interface.value"
   TextField "Line Label" at 0,0 size 267x40; Text 'Line:'
      Visibility <- "interface.animate.bg"
      Appearance <- "interface.animate.bg"
*)

(* ===== HMI "HMI_RT_1" =====

ScreenModuleEditorView "LED Row" 440x28
   TextField "tfLine" at 0,0 size 110x28; Text 'Text'
      Visibility <- "interface.tfLine.animate"
      Appearance <- "interface.tfLine.animate"
   TextField "tfTime" at 349,0 size 91x28; Text 'Text'
      Visibility <- "interface.tfTime.animate"
      Appearance <- "interface.tfTime.animate"
   TextField "tfDropZone" at 105,0 size 42x28; Text 'Text'
      Visibility <- "interface.tfDropZone.animate"
      Appearance <- "interface.tfDropZone.animate"
   TextField "tfSLPartNumber" at 146,0 size 209x28; Text 'Text'
      Visibility <- "interface.tfPartNumber.animateSL"
      Appearance <- "interface.tfPartNumber.animateSL"
   TextField "tfDLPartNumber" at 146,0 size 209x28; Text 'Text'
      Visibility <- "interface.tfPartNumber.animateDL"
      Appearance <- "interface.tfPartNumber.animateDL"
*)

(* ===== HMI "HMI_RT_1" =====
system functions are stored by id; their names below are inferred from use

ScreenModuleEditorView "IO Field: Timer" 137x50
   IOField "Allotted Time Entry Field" at 0,0 size 137x50; FormatPattern ???????
      on OnFinishInput: SetBit("Interface.inputFinished")
      Appearance <- "Interface.animate"
      Visibility <- "Interface.animate"
      ObjectEnable <- "Interface.animate"
      ProcessValue <- "Interface.value"
*)

(* ===== HMI "HMI_RT_1" =====
system functions are stored by id; their names below are inferred from use

ScreenModuleEditorView "IO Field: Double Width; Stacked" 414x50
   IOField "PN Entry Field" at 0,0 size 414x50; FormatPattern ????????????????????????????????????????
      on OnFinishInput: SetBit("Interface.inputFinished")
      Appearance <- "Interface.animate"
      Visibility <- "Interface.animate"
      ObjectEnable <- "Interface.animate"
      ProcessValue <- "Interface.value"
*)

(* ===== HMI "HMI_RT_1" =====
system functions are stored by id; their names below are inferred from use

ScreenModuleEditorView "Drop Zone Label" 240x40
   IOField "Drop Zone Entry" at 171,0 size 69x40; FormatPattern ??
      on OnFinishInput: SetBit("Interface.inputFinished")
      Appearance <- "Interface.animate.ioField"
      Visibility <- "Interface.animate.ioField"
      ProcessValue <- "Interface.value"
      ObjectEnable <- "Interface.animate.ioField"
   TextField "Drop Zone Label" at 0,0 size 240x40; Text 'Drop Zone:'
      Visibility <- "Interface.animate.bg"
      Appearance <- "Interface.animate.bg"
*)

(* ===== HMI "HMI_RT_1" =====
system functions are stored by id; their names below are inferred from use

ScreenModuleEditorView "PB: Station Comm Status (Text Label)" 205x65
   Button "Station Select" at 0,0 size 205x65; TextOff 'Text'
      on Press: function_b14e0dd5("Interface.actuate", 0)
      Appearance <- "Interface.animate"
      ObjectEnable <- "Interface.animate"
      Visibility <- "Interface.animate"
*)

(* ===== HMI "HMI_RT_1" =====
system functions are stored by id; their names below are inferred from use